// TIA Portal project "erronka5_talde2_v3" (V16)

(* hardware
DEVICE "S7-1200 station_1"  S7-1200 Station
   slot 0: "Rack_0"  S7-1200 Rack  Rack  V1.0
   slot 1: "PLC_1"  CPU 1215C AC/DC/Rly  6ES7 215-1BG40-0XB0  V4.2
*)

// ===== PLC "PLC_1"  CPU 1215C AC/DC/Rly =====

VAR_GLOBAL   // PLC tag table "Tabla de variables estándar"
   "M_VarTemporizador" AT %MD132 : Time;
   "SCA_A_Plus" AT %M120.1 : Bool;
   "IN_FC_C1" AT %I0.6 : Bool;
   "M_Et_59" AT %M51.1 : Bool;
   "M_Et_60" AT %M51.2 : Bool;
END_VAR

VAR_GLOBAL   // PLC tag table "VARS_SCADA>>PLC"
   "M_ConsignaCiclos" AT %MW168 : Int;
   "M_Balb_1_Act" AT %M20.3 : Bool;   // Lehenengo balbula aktibatzeko memoria, kontrol manuala dugunean.
   "M_Balb_2_Act" AT %M20.4 : Bool;   // Lehenengo balbula desaktibatzeko memoria, kontrol manuala dugunean.
   "M_Cil_Bultzatu" AT %M20.5 : Bool;   // Pieza bultzatzen duen zilindroaren aktibazioa.
   "M_Manual_Override" AT %M20.6 : Bool;
   "M_material_index" AT %MW172 : Int;
   "M_Var_Velocidad" AT %MD148 : Real;
   "M_Reset" AT %M165.0 : Bool;
END_VAR

VAR_GLOBAL   // PLC tag table "ETAPAK"
   "M_Et_20" AT %M20.0 : Bool;
   "M_Et_21" AT %M20.1 : Bool;
   "M_Et_30" AT %M30.0 : Bool;
   "M_Et_31" AT %M30.1 : Bool;
   "M_Et_40" AT %M40.0 : Bool;
   "M_Et_41" AT %M40.1 : Bool;
   "M_Et_100" AT %M100.0 : Bool;
   "M_Et_101" AT %M100.1 : Bool;
   "M_Et_50" AT %M50.0 : Bool;
   "M_Et_51" AT %M50.1 : Bool;
   "M_Et_52" AT %M50.2 : Bool;
   "M_Et_53" AT %M50.3 : Bool;
   "M_Et_54" AT %M50.4 : Bool;
   "M_Et_55" AT %M50.5 : Bool;
   "M_Et_56" AT %M50.6 : Bool;
   "M_Et_57" AT %M50.7 : Bool;
   "M_Et_58" AT %M51.0 : Bool;
   "M_Et_0" AT %M16.0 : Bool;
END_VAR

VAR_GLOBAL   // PLC tag table "VARS_PLC>>SCADA"
   "M_PisuaNorm" AT %MD124 : Real;
   "M_Num_Ciclos_Act" AT %MW170 : Int;
   "M_Status_Valv_1" AT %MW176 : Int;
   "M_Status_Valv_2" AT %MW178 : Int;
   "M_Status_Cil" AT %MW180 : Int;
END_VAR

VAR_GLOBAL   // PLC tag table "SARRERAK"
   "IN_Boton_Paro" AT %I1.0 : Bool;
   "IN_Pisua_Analog" AT %IW64 : Word;
   "IN_Martxa" AT %I0.0 : Bool;
   "IN_Tenperatura" AT %I0.1 : Bool;
   "IN_FC_A0" AT %I0.2 : Bool;
   "IN_FC_A1" AT %I0.3 : Bool;
   "IN_FC_B0" AT %I0.4 : Bool;
   "IN_FC_B1" AT %I0.5 : Bool;
   "IN_FC_C0" AT %I0.7 : Bool;
END_VAR

VAR_GLOBAL   // PLC tag table "IRTEERAK"
   "OUT_MotorON" AT %Q0.6 : Bool;
   "OUT_ConsignaVelocidad" AT %QW64 : Word;
   "OUT_A_plus" AT %Q0.0 : Bool;
   "OUT_A_minus" AT %Q0.1 : Bool;
   "OUT_B_plus" AT %Q0.2 : Bool;
   "OUT_B_minus" AT %Q0.3 : Bool;
   "OUT_C_plus" AT %Q0.4 : Bool;
   "OUT_Rele_Reg" AT %Q0.5 : Bool;
END_VAR

VAR_GLOBAL   // PLC tag table "MARKAK"
   "M_Velocidad_Norm" AT %MD164 : Real;
   "M_Peso_Ciclo" AT %MD120 : Real;
   "M_Pisua_KG" AT %MD128 : Real;
   "WEB_ERRORERAKO_MARKA" AT %MW174 : Int;
END_VAR

// folder: System blocks/Program resources

DATA_BLOCK "T1"   // DB1
{ S7_Optimized_Access := 'TRUE' }
AUTHOR : Simatic
FAMILY : IEC
NAME : IEC_TMR
VERSION : 1.0
// stored: InstanceOfName IEC_TIMER
"IEC_TIMER"
BEGIN
END_DATA_BLOCK

DATA_BLOCK "Temporizador motorea"   // DB2
{ S7_Optimized_Access := 'TRUE' }
AUTHOR : Simatic
FAMILY : IEC
NAME : IEC_TMR
VERSION : 1.0
// stored: InstanceOfName IEC_TIMER
"IEC_TIMER"
BEGIN
END_DATA_BLOCK

DATA_BLOCK "Denborak"   // DB3
{ S7_Optimized_Access := 'TRUE' }
VERSION : 0.1
   VAR
      materialen_denborak : Array[0..5] of Time;
   END_VAR
BEGIN
   materialen_denborak[0] := T#2S;
   materialen_denborak[1] := T#5S;
   materialen_denborak[2] := T#10S;
   materialen_denborak[3] := T#12S;
   materialen_denborak[4] := T#3S_500MS;
   materialen_denborak[5] := T#8S;
END_DATA_BLOCK

DATA_BLOCK "Abiadurak"   // DB4
{ S7_Optimized_Access := 'TRUE' }
VERSION : 0.1
   VAR
      Motorearen_abiadura : Array[0..5] of Real;
   END_VAR
BEGIN
   Motorearen_abiadura[0] := 40.0;
   Motorearen_abiadura[1] := 15.0;
   Motorearen_abiadura[2] := 30.0;
   Motorearen_abiadura[3] := 10.0;
   Motorearen_abiadura[4] := 40.0;
   Motorearen_abiadura[5] := 25.0;
END_DATA_BLOCK

DATA_BLOCK "IEC_Counter_0_DB_1"   // DB5
{ S7_Optimized_Access := 'TRUE' }
AUTHOR : Simatic
FAMILY : IEC
NAME : CNTR
VERSION : 1.0
// stored: InstanceOfName IEC_COUNTER
"IEC_COUNTER"
BEGIN
END_DATA_BLOCK

// folder: (top level)

FUNCTION "Zikloa" : Void   // FC1, LAD
{ S7_Optimized_Access := 'TRUE' }
VERSION : 0.1
BEGIN

REGION Network 1
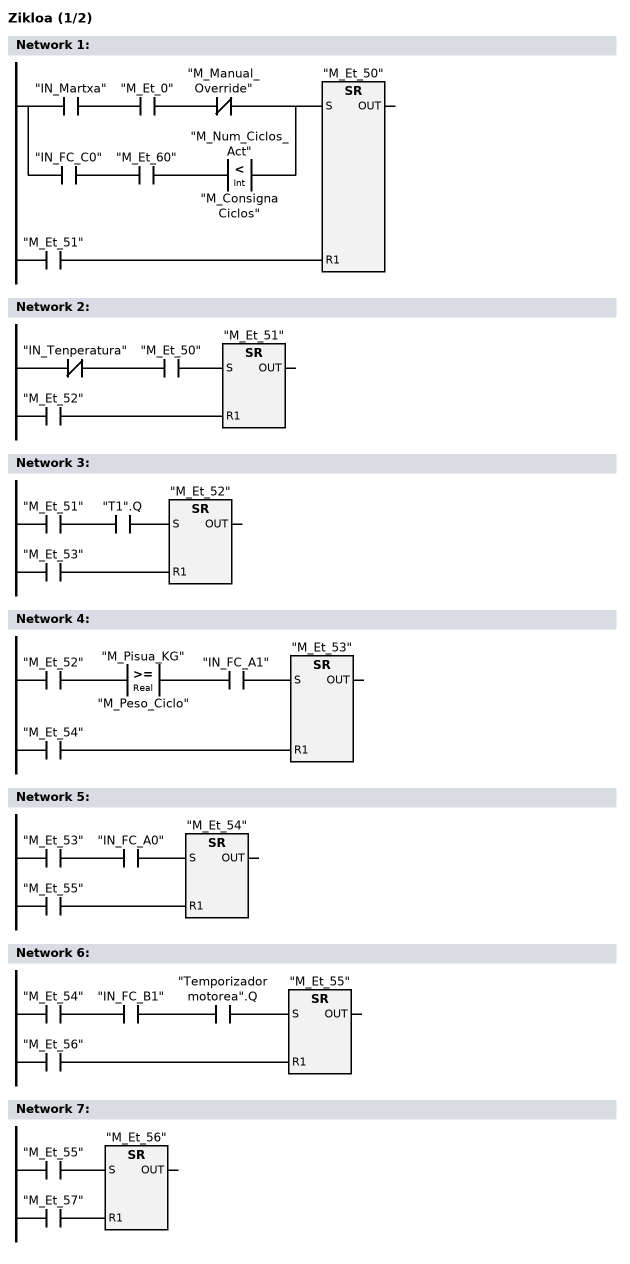
   RUNG wire#powerrail
      Contact( "IN_Martxa" )
      Contact( "M_Et_0" )
      I_Contact( "M_Manual_Override" )
      wire#w1
      S_SR(operand := "M_Et_50", r1 := wire#w2)
   END_RUNG
   RUNG wire#powerrail
      Contact( "IN_FC_C0" )
      Contact( "M_Et_60" )
      { S7_Templates := "SrcType := Int" } LT_Contact(in1 := "M_Num_Ciclos_Act", in2 := "M_ConsignaCiclos")
   END_RUNG wire#w1
   RUNG wire#powerrail
      Contact( "M_Et_51" )
   END_RUNG wire#w2
   // the same network as SCL:
   IF ("IN_Martxa" AND "M_Et_0" AND NOT "M_Manual_Override") OR ("IN_FC_C0" AND "M_Et_60" AND ("M_Num_Ciclos_Act" < "M_ConsignaCiclos")) THEN
       "M_Et_50" := TRUE;   // SR flip-flop
   END_IF;
   IF "M_Et_51" THEN "M_Et_50" := FALSE; END_IF;
END_REGION

REGION Network 2
   RUNG wire#powerrail
      I_Contact( "IN_Tenperatura" )
      Contact( "M_Et_50" )
      S_SR(operand := "M_Et_51", r1 := wire#w1)
   END_RUNG
   RUNG wire#powerrail
      Contact( "M_Et_52" )
   END_RUNG wire#w1
   // the same network as SCL:
   IF NOT "IN_Tenperatura" AND "M_Et_50" THEN
       "M_Et_51" := TRUE;   // SR flip-flop
   END_IF;
   IF "M_Et_52" THEN "M_Et_51" := FALSE; END_IF;
END_REGION

REGION Network 3
   RUNG wire#powerrail
      Contact( "M_Et_51" )
      Contact( "T1".Q )
      S_SR(operand := "M_Et_52", r1 := wire#w1)
   END_RUNG
   RUNG wire#powerrail
      Contact( "M_Et_53" )
   END_RUNG wire#w1
   // the same network as SCL:
   IF "M_Et_51" AND "T1".Q THEN
       "M_Et_52" := TRUE;   // SR flip-flop
   END_IF;
   IF "M_Et_53" THEN "M_Et_52" := FALSE; END_IF;
END_REGION

REGION Network 4
   RUNG wire#powerrail
      Contact( "M_Et_52" )
      { S7_Templates := "SrcType := Real" } GE_Contact(in1 := "M_Pisua_KG", in2 := "M_Peso_Ciclo")
      Contact( "IN_FC_A1" )
      S_SR(operand := "M_Et_53", r1 := wire#w1)
   END_RUNG
   RUNG wire#powerrail
      Contact( "M_Et_54" )
   END_RUNG wire#w1
   // the same network as SCL:
   IF "M_Et_52" AND ("M_Pisua_KG" >= "M_Peso_Ciclo") AND "IN_FC_A1" THEN
       "M_Et_53" := TRUE;   // SR flip-flop
   END_IF;
   IF "M_Et_54" THEN "M_Et_53" := FALSE; END_IF;
END_REGION

REGION Network 5
   RUNG wire#powerrail
      Contact( "M_Et_53" )
      Contact( "IN_FC_A0" )
      S_SR(operand := "M_Et_54", r1 := wire#w1)
   END_RUNG
   RUNG wire#powerrail
      Contact( "M_Et_55" )
   END_RUNG wire#w1
   // the same network as SCL:
   IF "M_Et_53" AND "IN_FC_A0" THEN
       "M_Et_54" := TRUE;   // SR flip-flop
   END_IF;
   IF "M_Et_55" THEN "M_Et_54" := FALSE; END_IF;
END_REGION

REGION Network 6
   RUNG wire#powerrail
      Contact( "M_Et_54" )
      Contact( "IN_FC_B1" )
      Contact( "Temporizador motorea".Q )
      S_SR(operand := "M_Et_55", r1 := wire#w1)
   END_RUNG
   RUNG wire#powerrail
      Contact( "M_Et_56" )
   END_RUNG wire#w1
   // the same network as SCL:
   IF "M_Et_54" AND "IN_FC_B1" AND "Temporizador motorea".Q THEN
       "M_Et_55" := TRUE;   // SR flip-flop
   END_IF;
   IF "M_Et_56" THEN "M_Et_55" := FALSE; END_IF;
END_REGION

REGION Network 7
   RUNG wire#powerrail
      Contact( "M_Et_55" )
      S_SR(operand := "M_Et_56", r1 := wire#w1)
   END_RUNG
   RUNG wire#powerrail
      Contact( "M_Et_57" )
   END_RUNG wire#w1
   // the same network as SCL:
   IF "M_Et_55" THEN
       "M_Et_56" := TRUE;   // SR flip-flop
   END_IF;
   IF "M_Et_57" THEN "M_Et_56" := FALSE; END_IF;
END_REGION

REGION Network 8
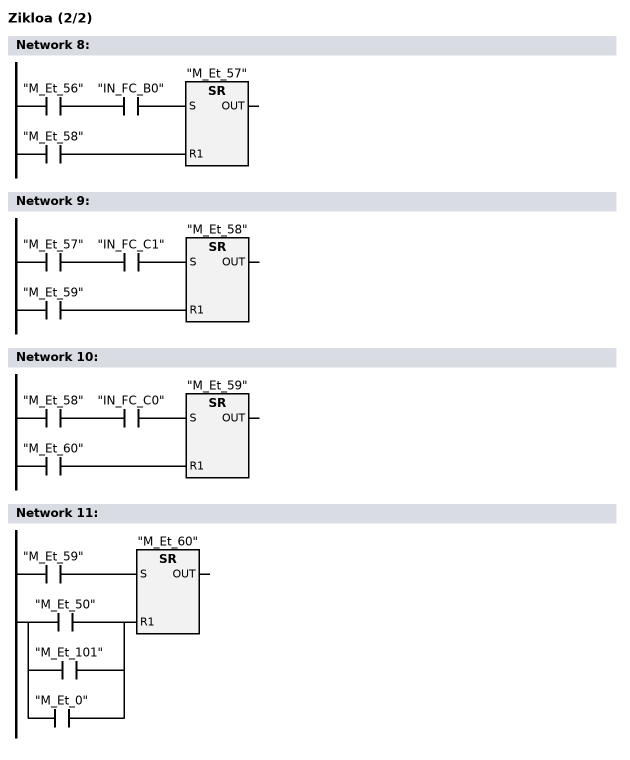
   RUNG wire#powerrail
      Contact( "M_Et_56" )
      Contact( "IN_FC_B0" )
      S_SR(operand := "M_Et_57", r1 := wire#w1)
   END_RUNG
   RUNG wire#powerrail
      Contact( "M_Et_58" )
   END_RUNG wire#w1
   // the same network as SCL:
   IF "M_Et_56" AND "IN_FC_B0" THEN
       "M_Et_57" := TRUE;   // SR flip-flop
   END_IF;
   IF "M_Et_58" THEN "M_Et_57" := FALSE; END_IF;
END_REGION

REGION Network 9
   RUNG wire#powerrail
      Contact( "M_Et_57" )
      Contact( "IN_FC_C1" )
      S_SR(operand := "M_Et_58", r1 := wire#w1)
   END_RUNG
   RUNG wire#powerrail
      Contact( "M_Et_59" )
   END_RUNG wire#w1
   // the same network as SCL:
   IF "M_Et_57" AND "IN_FC_C1" THEN
       "M_Et_58" := TRUE;   // SR flip-flop
   END_IF;
   IF "M_Et_59" THEN "M_Et_58" := FALSE; END_IF;
END_REGION

REGION Network 10
   RUNG wire#powerrail
      Contact( "M_Et_58" )
      Contact( "IN_FC_C0" )
      S_SR(operand := "M_Et_59", r1 := wire#w1)
   END_RUNG
   RUNG wire#powerrail
      Contact( "M_Et_60" )
   END_RUNG wire#w1
   // the same network as SCL:
   IF "M_Et_58" AND "IN_FC_C0" THEN
       "M_Et_59" := TRUE;   // SR flip-flop
   END_IF;
   IF "M_Et_60" THEN "M_Et_59" := FALSE; END_IF;
END_REGION

REGION Network 11
   RUNG wire#powerrail
      Contact( "M_Et_59" )
      S_SR(operand := "M_Et_60", r1 := wire#w1)
   END_RUNG
   RUNG wire#powerrail
      Contact( "M_Et_50" )
   END_RUNG wire#w1
   RUNG wire#powerrail
      Contact( "M_Et_101" )
   END_RUNG wire#w1
   RUNG wire#powerrail
      Contact( "M_Et_0" )
   END_RUNG wire#w1
   // the same network as SCL:
   IF "M_Et_59" THEN
       "M_Et_60" := TRUE;   // SR flip-flop
   END_IF;
   IF "M_Et_50" OR "M_Et_101" OR "M_Et_0" THEN "M_Et_60" := FALSE; END_IF;
END_REGION
END_FUNCTION

FUNCTION "Paro" : Void   // FC2, LAD
{ S7_Optimized_Access := 'TRUE' }
VERSION : 0.1
BEGIN

REGION Network 1
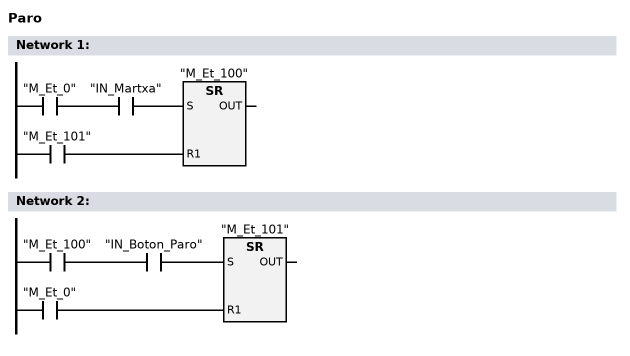
   RUNG wire#powerrail
      Contact( "M_Et_0" )
      Contact( "IN_Martxa" )
      S_SR(operand := "M_Et_100", r1 := wire#w1)
   END_RUNG
   RUNG wire#powerrail
      Contact( "M_Et_101" )
   END_RUNG wire#w1
   // the same network as SCL:
   IF "M_Et_0" AND "IN_Martxa" THEN
       "M_Et_100" := TRUE;   // SR flip-flop
   END_IF;
   IF "M_Et_101" THEN "M_Et_100" := FALSE; END_IF;
END_REGION

REGION Network 2
   RUNG wire#powerrail
      Contact( "M_Et_100" )
      Contact( "IN_Boton_Paro" )
      S_SR(operand := "M_Et_101", r1 := wire#w1)
   END_RUNG
   RUNG wire#powerrail
      Contact( "M_Et_0" )
   END_RUNG wire#w1
   // the same network as SCL:
   IF "M_Et_100" AND "IN_Boton_Paro" THEN
       "M_Et_101" := TRUE;   // SR flip-flop
   END_IF;
   IF "M_Et_0" THEN "M_Et_101" := FALSE; END_IF;
END_REGION
END_FUNCTION

FUNCTION "Akzioak" : Void   // FC3, LAD
{ S7_Optimized_Access := 'TRUE' }
VERSION : 0.1
BEGIN

REGION Network 1
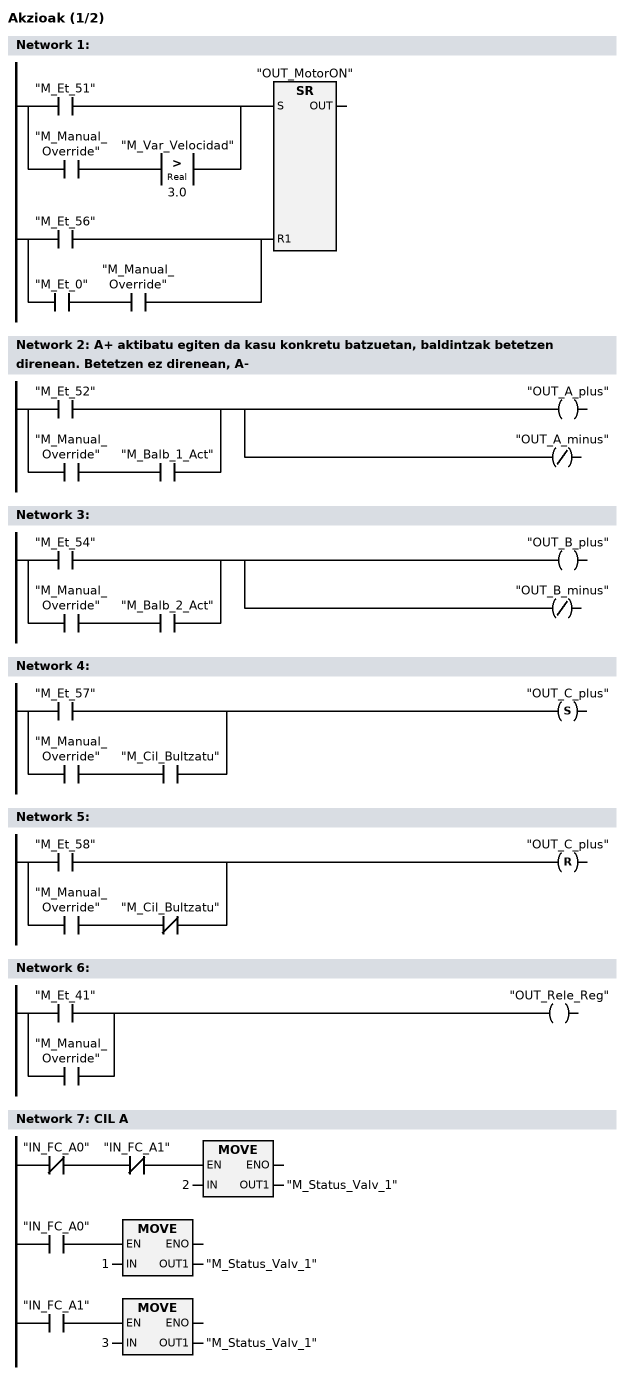
   RUNG wire#powerrail
      Contact( "M_Et_51" )
      wire#w1
      S_SR(operand := "OUT_MotorON", r1 := wire#w2)
   END_RUNG
   RUNG wire#powerrail
      Contact( "M_Manual_Override" )
      { S7_Templates := "SrcType := Real" } GT_Contact(in1 := "M_Var_Velocidad", in2 := 3.0)
   END_RUNG wire#w1
   RUNG wire#powerrail
      Contact( "M_Et_56" )
   END_RUNG wire#w2
   RUNG wire#powerrail
      Contact( "M_Et_0" )
      Contact( "M_Manual_Override" )
   END_RUNG wire#w2
   // the same network as SCL:
   IF "M_Et_51" OR ("M_Manual_Override" AND ("M_Var_Velocidad" > 3.0)) THEN
       "OUT_MotorON" := TRUE;   // SR flip-flop
   END_IF;
   IF "M_Et_56" OR ("M_Et_0" AND "M_Manual_Override") THEN "OUT_MotorON" := FALSE; END_IF;
END_REGION

REGION Network 2: A+ aktibatu egiten da kasu konkretu batzuetan, baldintzak betetzen direnean. Betetzen ez direnean, A-
   RUNG wire#powerrail
      Contact( "M_Et_52" )
      wire#w1
      Coil( "OUT_A_plus" )
   END_RUNG
   RUNG wire#powerrail
      Contact( "M_Manual_Override" )
      Contact( "M_Balb_1_Act" )
   END_RUNG wire#w1
   RUNG wire#w1
      I_Coil( "OUT_A_minus" )
   END_RUNG
   // the same network as SCL:
   "OUT_A_plus" := "M_Et_52" OR ("M_Manual_Override" AND "M_Balb_1_Act");
   "OUT_A_minus" := NOT "OUT_A_plus";
END_REGION

REGION Network 3
   RUNG wire#powerrail
      Contact( "M_Et_54" )
      wire#w1
      Coil( "OUT_B_plus" )
   END_RUNG
   RUNG wire#powerrail
      Contact( "M_Manual_Override" )
      Contact( "M_Balb_2_Act" )
   END_RUNG wire#w1
   RUNG wire#w1
      I_Coil( "OUT_B_minus" )
   END_RUNG
   // the same network as SCL:
   "OUT_B_plus" := "M_Et_54" OR ("M_Manual_Override" AND "M_Balb_2_Act");
   "OUT_B_minus" := NOT "OUT_B_plus";
END_REGION

REGION Network 4
   RUNG wire#powerrail
      Contact( "M_Et_57" )
      wire#w1
      S_Coil( "OUT_C_plus" )
   END_RUNG
   RUNG wire#powerrail
      Contact( "M_Manual_Override" )
      Contact( "M_Cil_Bultzatu" )
   END_RUNG wire#w1
   // the same network as SCL:
   IF "M_Et_57" OR ("M_Manual_Override" AND "M_Cil_Bultzatu") THEN "OUT_C_plus" := TRUE; END_IF;
END_REGION

REGION Network 5
   RUNG wire#powerrail
      Contact( "M_Et_58" )
      wire#w1
      R_Coil( "OUT_C_plus" )
   END_RUNG
   RUNG wire#powerrail
      Contact( "M_Manual_Override" )
      I_Contact( "M_Cil_Bultzatu" )
   END_RUNG wire#w1
   // the same network as SCL:
   IF "M_Et_58" OR ("M_Manual_Override" AND NOT "M_Cil_Bultzatu") THEN "OUT_C_plus" := FALSE; END_IF;
END_REGION

REGION Network 6
   RUNG wire#powerrail
      Contact( "M_Et_41" )
      wire#w1
      Coil( "OUT_Rele_Reg" )
   END_RUNG
   RUNG wire#powerrail
      Contact( "M_Manual_Override" )
   END_RUNG wire#w1
   // the same network as SCL:
   "OUT_Rele_Reg" := "M_Et_41" OR "M_Manual_Override";
END_REGION

REGION Network 7: CIL A
   RUNG wire#powerrail
      I_Contact( "IN_FC_A0" )
      I_Contact( "IN_FC_A1" )
      Move(in := 2, out1 => "M_Status_Valv_1")
   END_RUNG
   RUNG wire#powerrail
      Contact( "IN_FC_A0" )
      Move(in := 1, out1 => "M_Status_Valv_1")
   END_RUNG
   RUNG wire#powerrail
      Contact( "IN_FC_A1" )
      Move(in := 3, out1 => "M_Status_Valv_1")
   END_RUNG
   // the same network as SCL:
   IF NOT "IN_FC_A0" AND NOT "IN_FC_A1" THEN "M_Status_Valv_1" := 2; END_IF;
   IF "IN_FC_A0" THEN "M_Status_Valv_1" := 1; END_IF;
   IF "IN_FC_A1" THEN "M_Status_Valv_1" := 3; END_IF;
END_REGION

REGION Network 8: CIL B
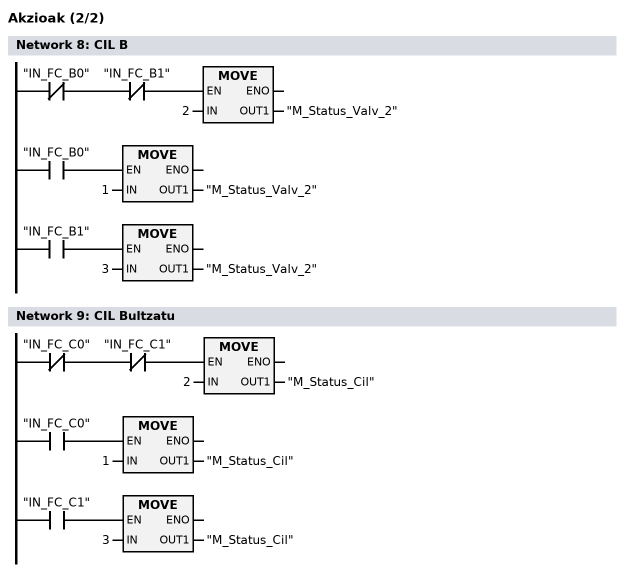
   RUNG wire#powerrail
      I_Contact( "IN_FC_B0" )
      I_Contact( "IN_FC_B1" )
      Move(in := 2, out1 => "M_Status_Valv_2")
   END_RUNG
   RUNG wire#powerrail
      Contact( "IN_FC_B0" )
      Move(in := 1, out1 => "M_Status_Valv_2")
   END_RUNG
   RUNG wire#powerrail
      Contact( "IN_FC_B1" )
      Move(in := 3, out1 => "M_Status_Valv_2")
   END_RUNG
   // the same network as SCL:
   IF NOT "IN_FC_B0" AND NOT "IN_FC_B1" THEN "M_Status_Valv_2" := 2; END_IF;
   IF "IN_FC_B0" THEN "M_Status_Valv_2" := 1; END_IF;
   IF "IN_FC_B1" THEN "M_Status_Valv_2" := 3; END_IF;
END_REGION

REGION Network 9: CIL Bultzatu
   RUNG wire#powerrail
      I_Contact( "IN_FC_C0" )
      I_Contact( "IN_FC_C1" )
      Move(in := 2, out1 => "M_Status_Cil")
   END_RUNG
   RUNG wire#powerrail
      Contact( "IN_FC_C0" )
      Move(in := 1, out1 => "M_Status_Cil")
   END_RUNG
   RUNG wire#powerrail
      Contact( "IN_FC_C1" )
      Move(in := 3, out1 => "M_Status_Cil")
   END_RUNG
   // the same network as SCL:
   IF NOT "IN_FC_C0" AND NOT "IN_FC_C1" THEN "M_Status_Cil" := 2; END_IF;
   IF "IN_FC_C0" THEN "M_Status_Cil" := 1; END_IF;
   IF "IN_FC_C1" THEN "M_Status_Cil" := 3; END_IF;
END_REGION
END_FUNCTION

FUNCTION "Temporizadoreak" : Void   // FC4, LAD
{ S7_Optimized_Access := 'TRUE' }
VERSION : 0.1
BEGIN

REGION Network 1
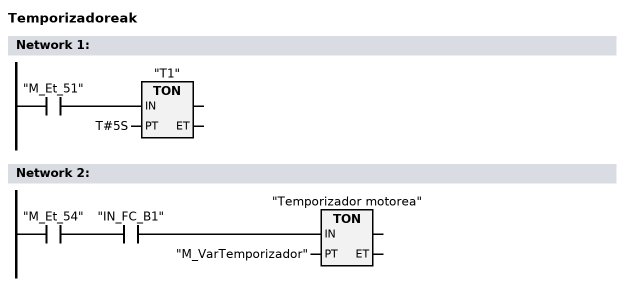
   "T1".TON(IN := "M_Et_51", PT := T#5S);
END_REGION

REGION Network 2
   "Temporizador motorea".TON(IN := "M_Et_54" AND "IN_FC_B1", PT := "M_VarTemporizador");
END_REGION
END_FUNCTION

FUNCTION "escalado" : Void   // FC5, LAD
{ S7_Optimized_Access := 'TRUE' }
VERSION : 0.1
BEGIN

REGION Network 1
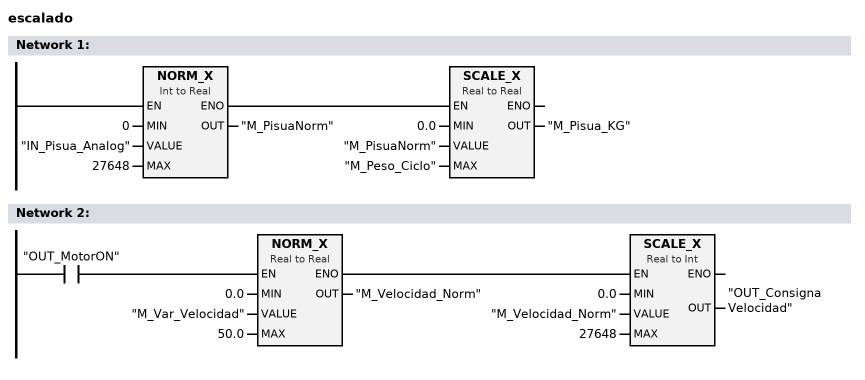
   RUNG wire#powerrail
      { S7_Templates := "[SrcType := Int, DestType := Real]" } Normalize(min := 0, value := "IN_Pisua_Analog", max := 27648, out => "M_PisuaNorm")
      { S7_Templates := "[SrcType := Real, DestType := Real]" } Scale(min := 0.0, value := "M_PisuaNorm", max := "M_Peso_Ciclo", out => "M_Pisua_KG")
   END_RUNG
   // the same network as SCL:
   "M_PisuaNorm" := NORM_X(MIN := 0, VALUE := "IN_Pisua_Analog", MAX := 27648);
   "M_Pisua_KG" := SCALE_X(MIN := 0.0, VALUE := "M_PisuaNorm", MAX := "M_Peso_Ciclo");
END_REGION

REGION Network 2
   RUNG wire#powerrail
      Contact( "OUT_MotorON" )
      { S7_Templates := "[SrcType := Real, DestType := Real]" } Normalize(min := 0.0, value := "M_Var_Velocidad", max := 50.0, out => "M_Velocidad_Norm")
      { S7_Templates := "[SrcType := Real, DestType := Int]" } Scale(min := 0.0, value := "M_Velocidad_Norm", max := 27648, out => "OUT_ConsignaVelocidad")
   END_RUNG
   // the same network as SCL:
   IF "OUT_MotorON" THEN
       "M_Velocidad_Norm" := NORM_X(MIN := 0.0, VALUE := "M_Var_Velocidad", MAX := 50.0);
       "OUT_ConsignaVelocidad" := SCALE_X(MIN := 0.0, VALUE := "M_Velocidad_Norm", MAX := 27648);
   END_IF;
END_REGION
END_FUNCTION

FUNCTION "Ziklo berogailua" : Void   // FC6, LAD
{ S7_Optimized_Access := 'TRUE' }
VERSION : 0.1
BEGIN

REGION Network 1
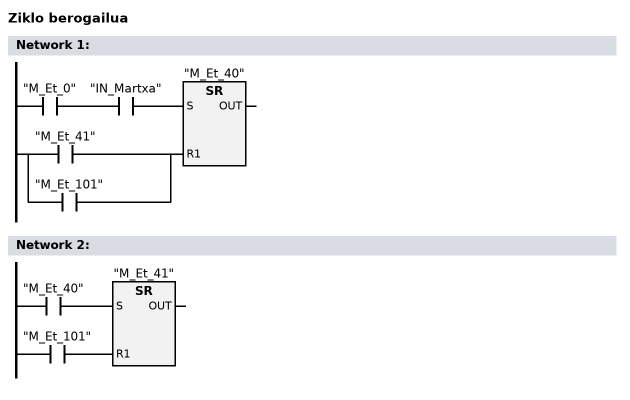
   RUNG wire#powerrail
      Contact( "M_Et_0" )
      Contact( "IN_Martxa" )
      S_SR(operand := "M_Et_40", r1 := wire#w1)
   END_RUNG
   RUNG wire#powerrail
      Contact( "M_Et_41" )
   END_RUNG wire#w1
   RUNG wire#powerrail
      Contact( "M_Et_101" )
   END_RUNG wire#w1
   // the same network as SCL:
   IF "M_Et_0" AND "IN_Martxa" THEN
       "M_Et_40" := TRUE;   // SR flip-flop
   END_IF;
   IF "M_Et_41" OR "M_Et_101" THEN "M_Et_40" := FALSE; END_IF;
END_REGION

REGION Network 2
   RUNG wire#powerrail
      Contact( "M_Et_40" )
      S_SR(operand := "M_Et_41", r1 := wire#w1)
   END_RUNG
   RUNG wire#powerrail
      Contact( "M_Et_101" )
   END_RUNG wire#w1
   // the same network as SCL:
   IF "M_Et_40" THEN
       "M_Et_41" := TRUE;   // SR flip-flop
   END_IF;
   IF "M_Et_101" THEN "M_Et_41" := FALSE; END_IF;
END_REGION
END_FUNCTION

FUNCTION "VariablesCiclo" : Void   // FC7, LAD
{ S7_Optimized_Access := 'TRUE' }
VERSION : 0.1
BEGIN

REGION Network 1
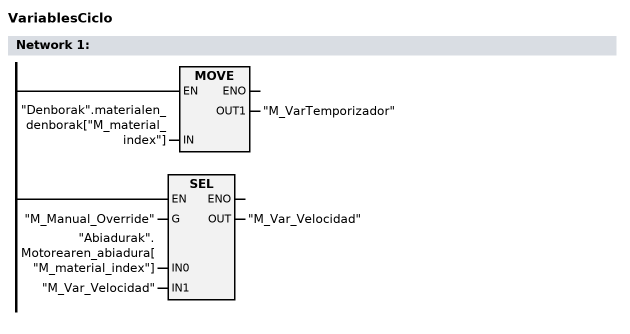
   "M_VarTemporizador" := "Denborak".materialen_denborak["M_material_index"];
   "M_Var_Velocidad" := SEL(G := "M_Manual_Override", IN0 := "Abiadurak".Motorearen_abiadura["M_material_index"], IN1 := "M_Var_Velocidad");
END_REGION
END_FUNCTION

FUNCTION "Contador" : Void   // FC10, LAD
{ S7_Optimized_Access := 'TRUE' }
VERSION : 0.1
BEGIN

REGION Network 1
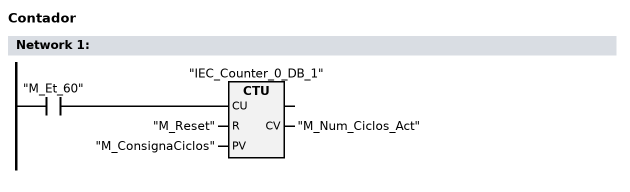
   "IEC_Counter_0_DB_1".CTU(CU := "M_Et_60", R := "M_Reset", PV := "M_ConsignaCiclos", CV => "M_Num_Ciclos_Act");
END_REGION
END_FUNCTION

ORGANIZATION_BLOCK "Main"   // OB1, LAD, ProgramCycle
TITLE = "Main Program Sweep (Cycle)"
{ S7_Optimized_Access := 'TRUE' }
VERSION : 0.1
   VAR_INPUT
      Initial_Call : Bool;   // Initial call of this OB
      Remanence : Bool;   // =True, if remanent data are available
   END_VAR
BEGIN

REGION Network 1
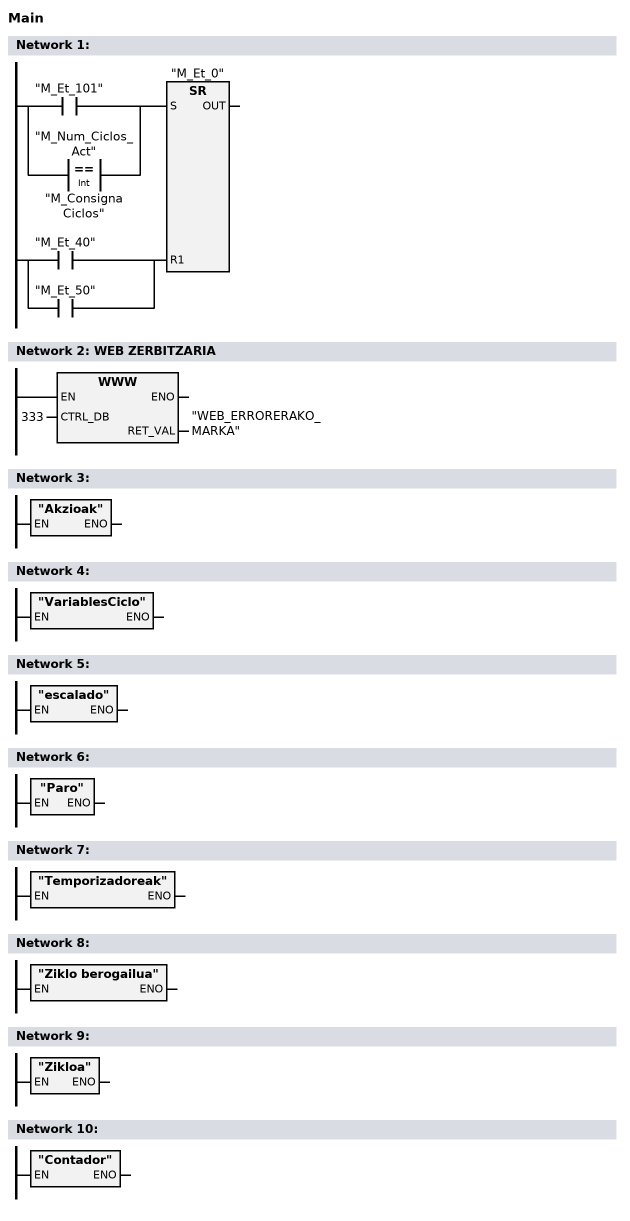
   RUNG wire#powerrail
      Contact( "M_Et_101" )
      wire#w1
      S_SR(operand := "M_Et_0", r1 := wire#w2)
   END_RUNG
   RUNG wire#powerrail
      { S7_Templates := "SrcType := Int" } EQ_Contact(in1 := "M_Num_Ciclos_Act", in2 := "M_ConsignaCiclos")
   END_RUNG wire#w1
   RUNG wire#powerrail
      Contact( "M_Et_40" )
   END_RUNG wire#w2
   RUNG wire#powerrail
      Contact( "M_Et_50" )
   END_RUNG wire#w2
   // the same network as SCL:
   IF "M_Et_101" OR ("M_Num_Ciclos_Act" = "M_ConsignaCiclos") THEN
       "M_Et_0" := TRUE;   // SR flip-flop
   END_IF;
   IF "M_Et_40" OR "M_Et_50" THEN "M_Et_0" := FALSE; END_IF;
END_REGION

REGION Network 2: WEB ZERBITZARIA
   "WEB_ERRORERAKO_MARKA" := WWW(CTRL_DB := 333);
END_REGION

REGION Network 3
   RUNG wire#powerrail
      "Akzioak"()
   END_RUNG
   // the same network as SCL:
   "Akzioak"();
END_REGION

REGION Network 4
   RUNG wire#powerrail
      "VariablesCiclo"()
   END_RUNG
   // the same network as SCL:
   "VariablesCiclo"();
END_REGION

REGION Network 5
   RUNG wire#powerrail
      "escalado"()
   END_RUNG
   // the same network as SCL:
   "escalado"();
END_REGION

REGION Network 6
   RUNG wire#powerrail
      "Paro"()
   END_RUNG
   // the same network as SCL:
   "Paro"();
END_REGION

REGION Network 7
   RUNG wire#powerrail
      "Temporizadoreak"()
   END_RUNG
   // the same network as SCL:
   "Temporizadoreak"();
END_REGION

REGION Network 8
   RUNG wire#powerrail
      "Ziklo berogailua"()
   END_RUNG
   // the same network as SCL:
   "Ziklo berogailua"();
END_REGION

REGION Network 9
   RUNG wire#powerrail
      "Zikloa"()
   END_RUNG
   // the same network as SCL:
   "Zikloa"();
END_REGION

REGION Network 10
   RUNG wire#powerrail
      "Contador"()
   END_RUNG
   // the same network as SCL:
   "Contador"();
END_REGION
END_ORGANIZATION_BLOCK

ORGANIZATION_BLOCK "Startup"   // OB100, LAD, Startup
TITLE = "Complete Restart"
{ S7_Optimized_Access := 'TRUE' }
VERSION : 0.1
   VAR_INPUT
      LostRetentive : Bool;   // True if retentive data are lost
      LostRTC : Bool;   // True if date and time are lost
   END_VAR
BEGIN

REGION Network 1
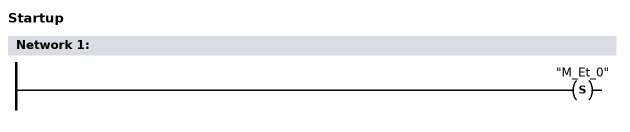
   RUNG wire#powerrail
      S_Coil( "M_Et_0" )
   END_RUNG
   // the same network as SCL:
   "M_Et_0" := TRUE;
END_REGION
END_ORGANIZATION_BLOCK